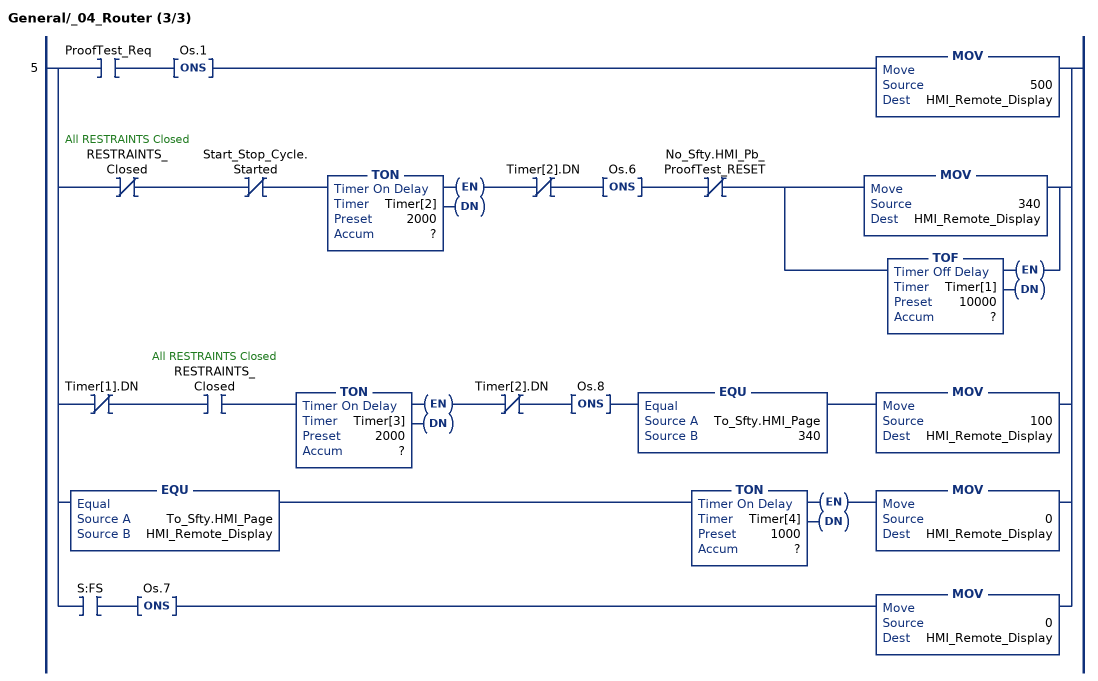
   5: [XIC(ProofTest_Req) ONS(Os.1) MOV(500,HMI_Remote_Display) ,XIO(RESTRAINTS_Closed) XIO(Start_Stop_Cycle.Started) TON(Timer[2],?,?) XIO(Timer[2].DN) ONS(Os.6) XIO(No_Sfty.HMI_Pb_ProofTest_RESET) [MOV(340,HMI_Remote_Display) ,TOF(Timer[1],?,?) ] ,XIO(Timer[1].DN) XIC(RESTRAINTS_Closed) TON(Timer[3],?,?) XIO(Timer[2].DN) ONS(Os.8) EQU(To_Sfty.HMI_Page,340) MOV(100,HMI_Remote_Display) ,EQU(To_Sfty.HMI_Page,HMI_Remote_Display) TON(Timer[4],?,?) MOV(0,HMI_Remote_Display) ,XIC(S:FS) ONS(Os.7) MOV(0,HMI_Remote_Display) ];
END_ROUTINE

ROUTINE _05_Miscellany   (* ladder *)
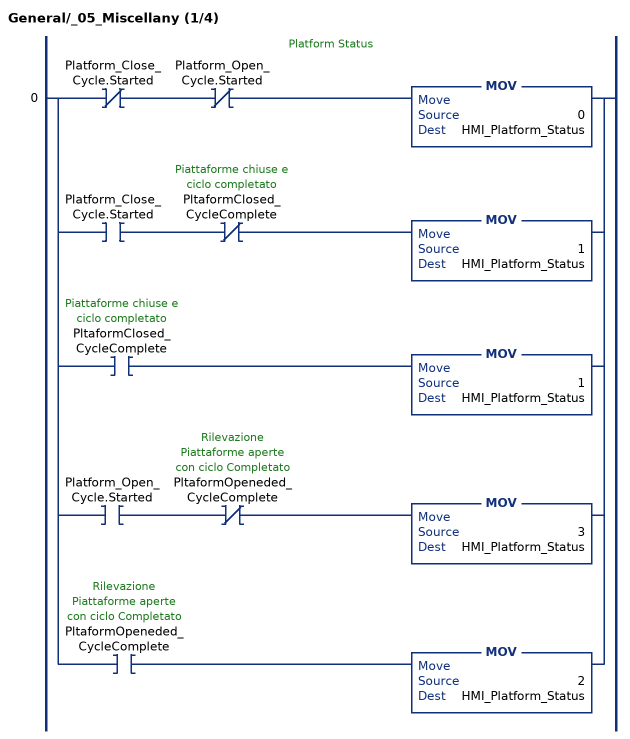
   // Platform Status
   0: [XIO(Platform_Close_Cycle.Started) XIO(Platform_Open_Cycle.Started) MOV(0,HMI_Platform_Status) ,XIC(Platform_Close_Cycle.Started) XIO(PltaformClosed_CycleComplete) MOV(1,HMI_Platform_Status) ,XIC(PltaformClosed_CycleComplete) MOV(1,HMI_Platform_Status) ,XIC(Platform_Open_Cycle.Started) XIO(PltaformOpeneded_CycleComplete) MOV(3,HMI_Platform_Status) ,XIC(PltaformOpeneded_CycleComplete) MOV(2,HMI_Platform_Status) ];
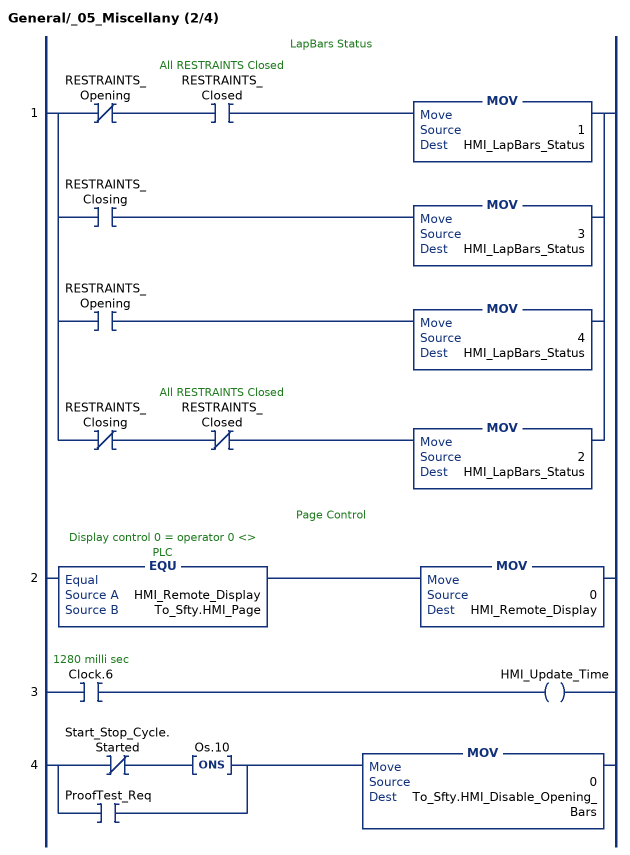
   // LapBars Status
   1: [XIO(RESTRAINTS_Opening) XIC(RESTRAINTS_Closed) MOV(1,HMI_LapBars_Status) ,XIC(RESTRAINTS_Closing) MOV(3,HMI_LapBars_Status) ,XIC(RESTRAINTS_Opening) MOV(4,HMI_LapBars_Status) ,XIO(RESTRAINTS_Closing) XIO(RESTRAINTS_Closed) MOV(2,HMI_LapBars_Status) ];
   // Page Control
   2: EQU(HMI_Remote_Display,To_Sfty.HMI_Page)MOV(0,HMI_Remote_Display);
   3: XIC(Clock.6)OTE(HMI_Update_Time);
   4: [XIO(Start_Stop_Cycle.Started) ONS(Os.10) ,XIC(ProofTest_Req) ]MOV(0,To_Sfty.HMI_Disable_Opening_Bars);
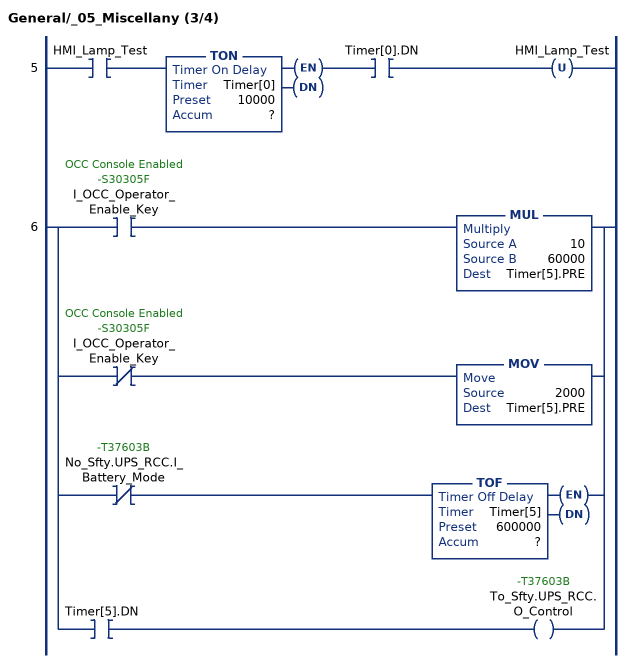
   5: XIC(HMI_Lamp_Test)TON(Timer[0],?,?)XIC(Timer[0].DN)OTU(HMI_Lamp_Test);
   6: [XIC(I_OCC_Operator_Enable_Key) MUL(10,60000,Timer[5].PRE) ,XIO(I_OCC_Operator_Enable_Key) MOV(2000,Timer[5].PRE) ,XIO(No_Sfty.UPS_RCC.I_Battery_Mode) TOF(Timer[5],?,?) ,XIC(Timer[5].DN) OTE(To_Sfty.UPS_RCC.O_Control) ];
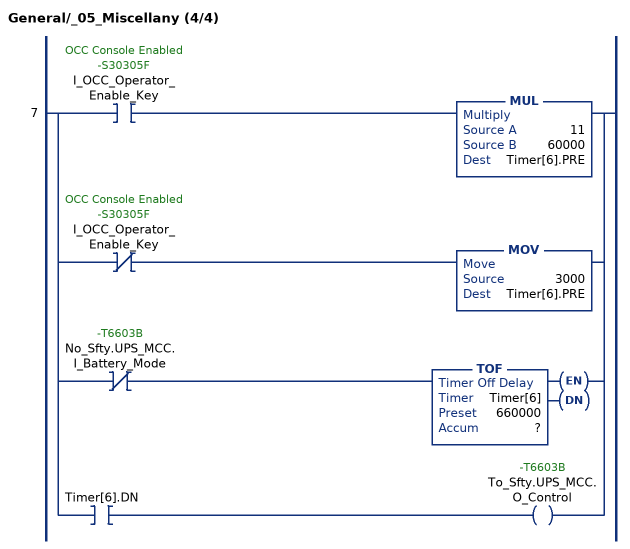
   7: [XIC(I_OCC_Operator_Enable_Key) MUL(11,60000,Timer[6].PRE) ,XIO(I_OCC_Operator_Enable_Key) MOV(3000,Timer[6].PRE) ,XIO(No_Sfty.UPS_MCC.I_Battery_Mode) TOF(Timer[6],?,?) ,XIC(Timer[6].DN) OTE(To_Sfty.UPS_MCC.O_Control) ];
END_ROUTINE

ROUTINE _06_HMI_Angle_Conversion   (* function block diagram *)
   SHEET 1
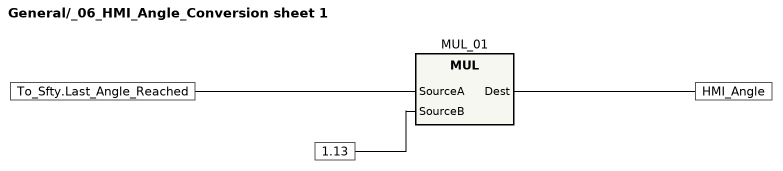
   MUL_01 : MUL(SourceA := To_Sfty.Last_Angle_Reached, SourceB := 1.13);
   HMI_Angle := MUL_01.Dest;
END_ROUTINE

ROUTINE _99_Statistics   (* ladder *)
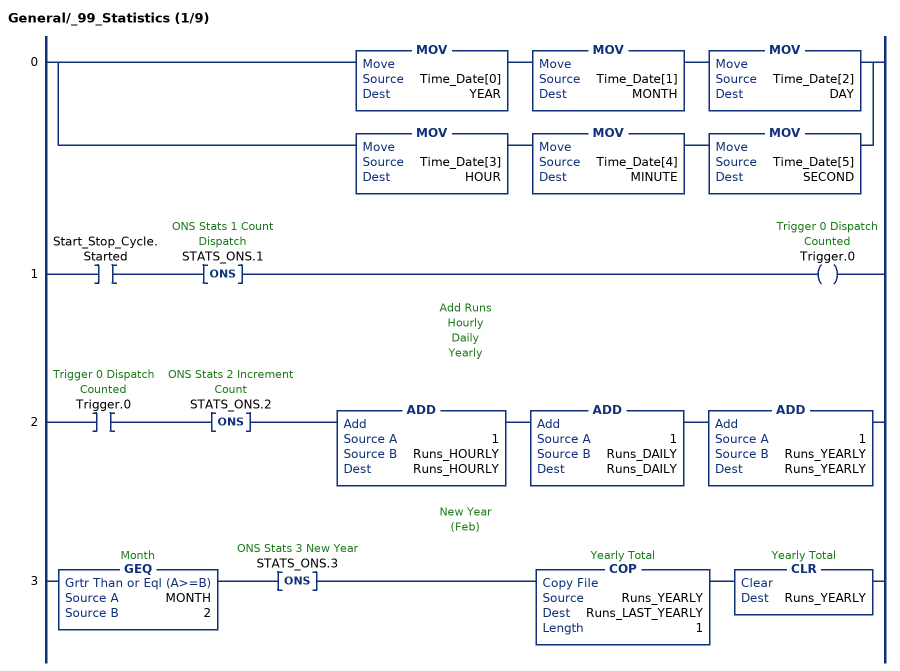
   0: [MOV(Time_Date[0],YEAR) MOV(Time_Date[1],MONTH) MOV(Time_Date[2],DAY) ,MOV(Time_Date[3],HOUR) MOV(Time_Date[4],MINUTE) MOV(Time_Date[5],SECOND) ];
   1: XIC(Start_Stop_Cycle.Started)ONS(STATS_ONS.1)OTE(Trigger.0);
   // Add Runs
   // Hourly
   // Daily
   // Yearly
   2: XIC(Trigger.0)ONS(STATS_ONS.2)ADD(1,Runs_HOURLY,Runs_HOURLY)ADD(1,Runs_DAILY,Runs_DAILY)ADD(1,Runs_YEARLY,Runs_YEARLY);
   // New Year
   // (Feb)
   3: GEQ(MONTH,2)ONS(STATS_ONS.3)COP(Runs_YEARLY,Runs_LAST_YEARLY,1)CLR(Runs_YEARLY);
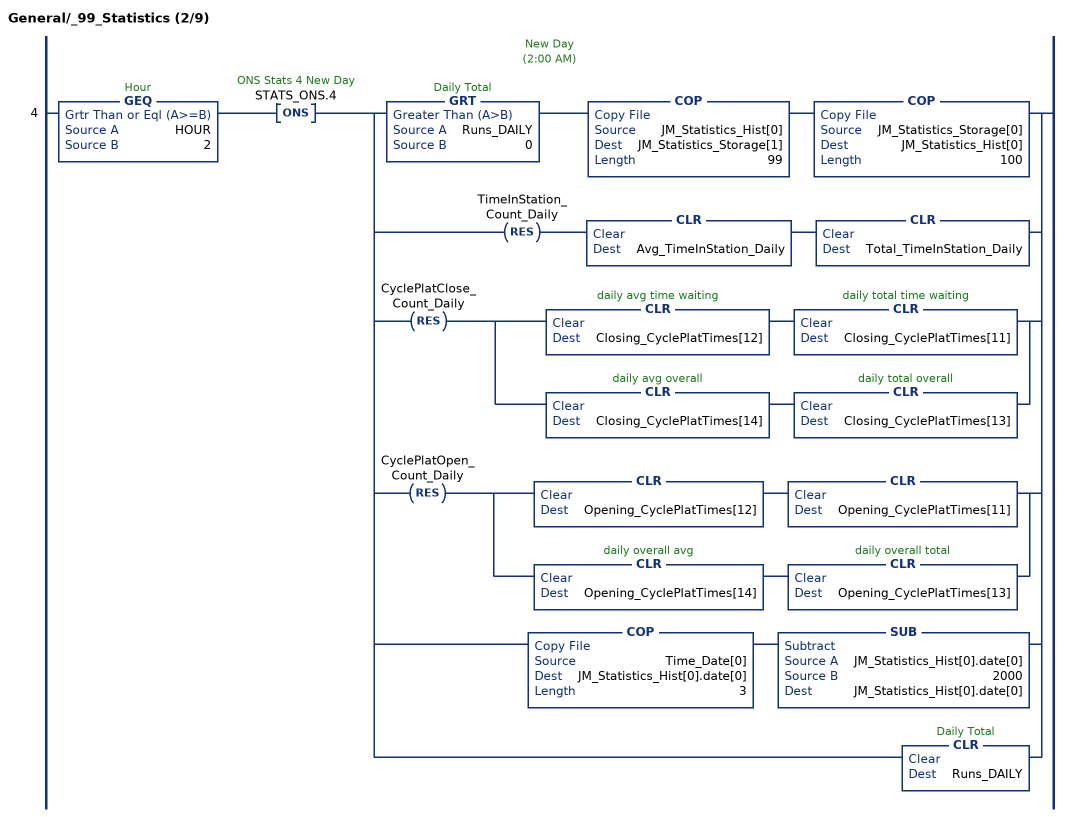
   // New Day
   // (2:00 AM)
   4: GEQ(HOUR,2)ONS(STATS_ONS.4)[[GRT(Runs_DAILY,0) COP(JM_Statistics_Hist[0],JM_Statistics_Storage[1],99) COP(JM_Statistics_Storage[0],JM_Statistics_Hist[0],100) ,RES(TimeInStation_Count_Daily) CLR(Avg_TimeInStation_Daily) CLR(Total_TimeInStation_Daily) ,RES(CyclePlatClose_Count_Daily) [CLR(Closing_CyclePlatTimes[12]) CLR(Closing_CyclePlatTimes[11]) ,CLR(Closing_CyclePlatTimes[14]) CLR(Closing_CyclePlatTimes[13]) ] ,RES(CyclePlatOpen_Count_Daily) [CLR(Opening_CyclePlatTimes[12]) CLR(Opening_CyclePlatTimes[11]) ,CLR(Opening_CyclePlatTimes[14]) CLR(Opening_CyclePlatTimes[13]) ] ,COP(Time_Date[0],JM_Statistics_Hist[0].date[0],3) SUB(JM_Statistics_Hist[0].date[0],2000,JM_Statistics_Hist[0].date[0]) ] ,CLR(Runs_DAILY) ];
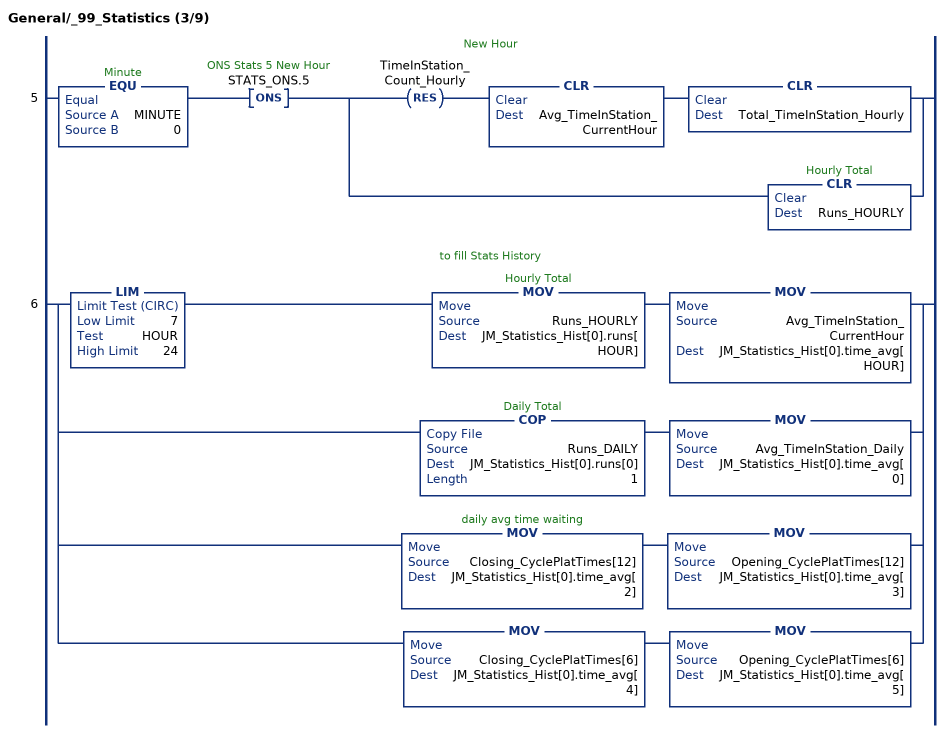
   // New Hour
   5: EQU(MINUTE,0)ONS(STATS_ONS.5)[RES(TimeInStation_Count_Hourly) CLR(Avg_TimeInStation_CurrentHour) CLR(Total_TimeInStation_Hourly) ,CLR(Runs_HOURLY) ];
   // to fill Stats History
   6: [LIM(7,HOUR,24) MOV(Runs_HOURLY,JM_Statistics_Hist[0].runs[HOUR]) MOV(Avg_TimeInStation_CurrentHour,JM_Statistics_Hist[0].time_avg[HOUR]) ,COP(Runs_DAILY,JM_Statistics_Hist[0].runs[0],1) MOV(Avg_TimeInStation_Daily,JM_Statistics_Hist[0].time_avg[0]) ,[MOV(Closing_CyclePlatTimes[12],JM_Statistics_Hist[0].time_avg[2]) MOV(Opening_CyclePlatTimes[12],JM_Statistics_Hist[0].time_avg[3]) ,MOV(Closing_CyclePlatTimes[6],JM_Statistics_Hist[0].time_avg[4]) MOV(Opening_CyclePlatTimes[6],JM_Statistics_Hist[0].time_avg[5]) ] ];
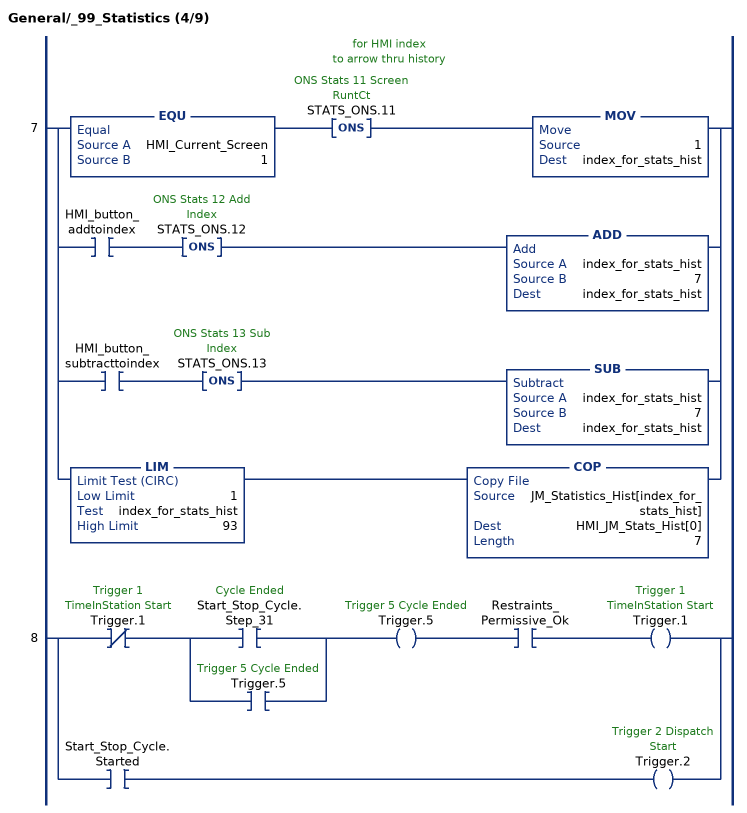
   // for HMI index
   // to arrow thru history
   7: [EQU(HMI_Current_Screen,1) ONS(STATS_ONS.11) MOV(1,index_for_stats_hist) ,[XIC(HMI_button_addtoindex) ONS(STATS_ONS.12) ADD(index_for_stats_hist,7,index_for_stats_hist) ,XIC(HMI_button_subtracttoindex) ONS(STATS_ONS.13) SUB(index_for_stats_hist,7,index_for_stats_hist) ] ,LIM(1,index_for_stats_hist,93) COP(JM_Statistics_Hist[index_for_stats_hist],HMI_JM_Stats_Hist[0],7) ];
   8: [XIO(Trigger.1) [XIC(Start_Stop_Cycle.Step_31) ,XIC(Trigger.5) ] OTE(Trigger.5) XIC(Restraints_Permissive_Ok) OTE(Trigger.1) ,XIC(Start_Stop_Cycle.Started) OTE(Trigger.2) ];
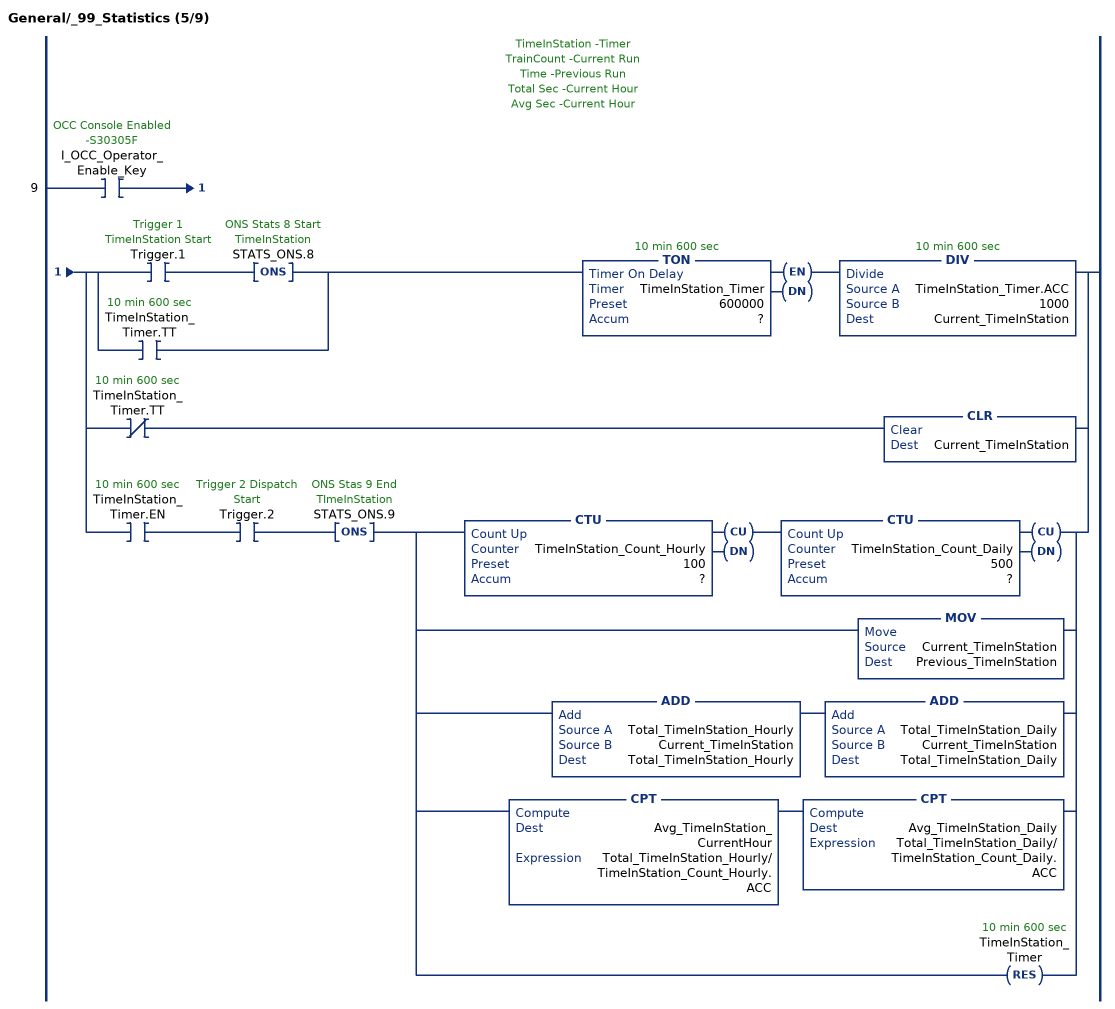
   // TimeInStation -Timer
   // TrainCount -Current Run
   // Time -Previous Run
   // Total Sec -Current Hour
   // Avg Sec -Current Hour
   9: XIC(I_OCC_Operator_Enable_Key)[[XIC(Trigger.1) ONS(STATS_ONS.8) ,XIC(TimeInStation_Timer.TT) ] TON(TimeInStation_Timer,?,?) DIV(TimeInStation_Timer.ACC,1000,Current_TimeInStation) ,XIO(TimeInStation_Timer.TT) CLR(Current_TimeInStation) ,XIC(TimeInStation_Timer.EN) XIC(Trigger.2) ONS(STATS_ONS.9) [CTU(TimeInStation_Count_Hourly,?,?) CTU(TimeInStation_Count_Daily,?,?) ,MOV(Current_TimeInStation,Previous_TimeInStation) ,ADD(Total_TimeInStation_Hourly,Current_TimeInStation,Total_TimeInStation_Hourly) ADD(Total_TimeInStation_Daily,Current_TimeInStation,Total_TimeInStation_Daily) ,CPT(Avg_TimeInStation_CurrentHour,Total_TimeInStation_Hourly/TimeInStation_Count_Hourly.ACC) CPT(Avg_TimeInStation_Daily,Total_TimeInStation_Daily/TimeInStation_Count_Daily.ACC) ,RES(TimeInStation_Timer) ] ];
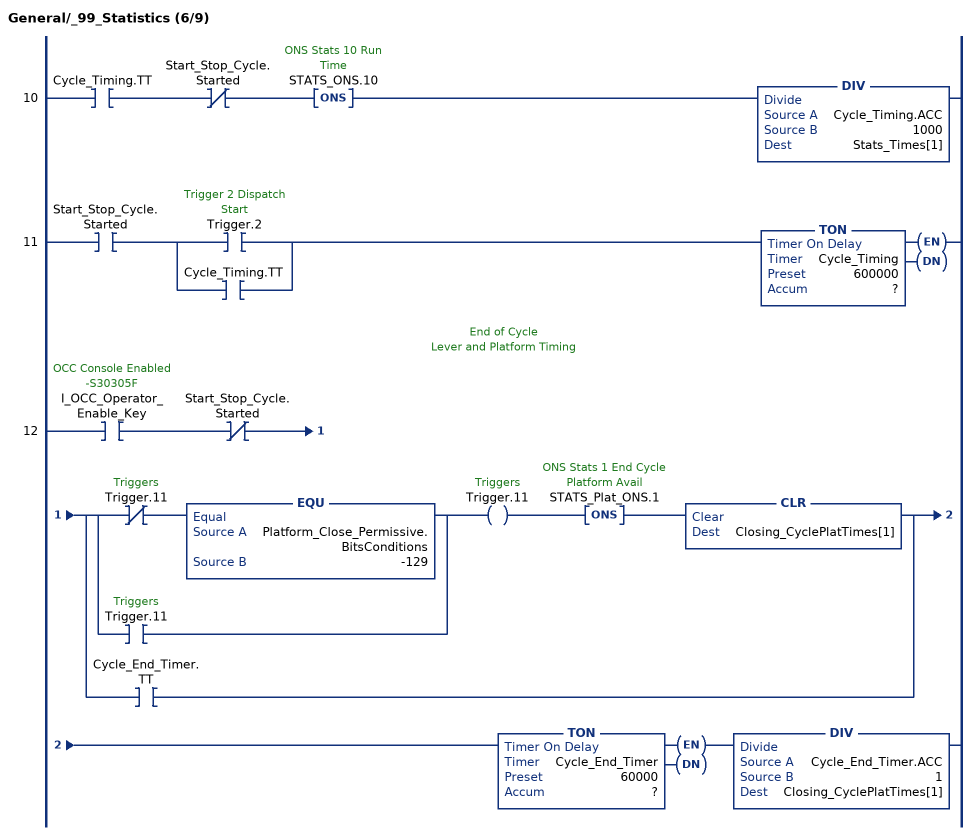
   10: XIC(Cycle_Timing.TT)XIO(Start_Stop_Cycle.Started)ONS(STATS_ONS.10)DIV(Cycle_Timing.ACC,1000,Stats_Times[1]);
   11: XIC(Start_Stop_Cycle.Started)[XIC(Trigger.2) ,XIC(Cycle_Timing.TT) ]TON(Cycle_Timing,?,?);
   // End of Cycle
   // Lever and Platform Timing
   12: XIC(I_OCC_Operator_Enable_Key)XIO(Start_Stop_Cycle.Started)[[XIO(Trigger.11) EQU(Platform_Close_Permissive.BitsConditions,-129) ,XIC(Trigger.11) ] OTE(Trigger.11) ONS(STATS_Plat_ONS.1) CLR(Closing_CyclePlatTimes[1]) ,XIC(Cycle_End_Timer.TT) ]TON(Cycle_End_Timer,?,?)DIV(Cycle_End_Timer.ACC,1,Closing_CyclePlatTimes[1]);
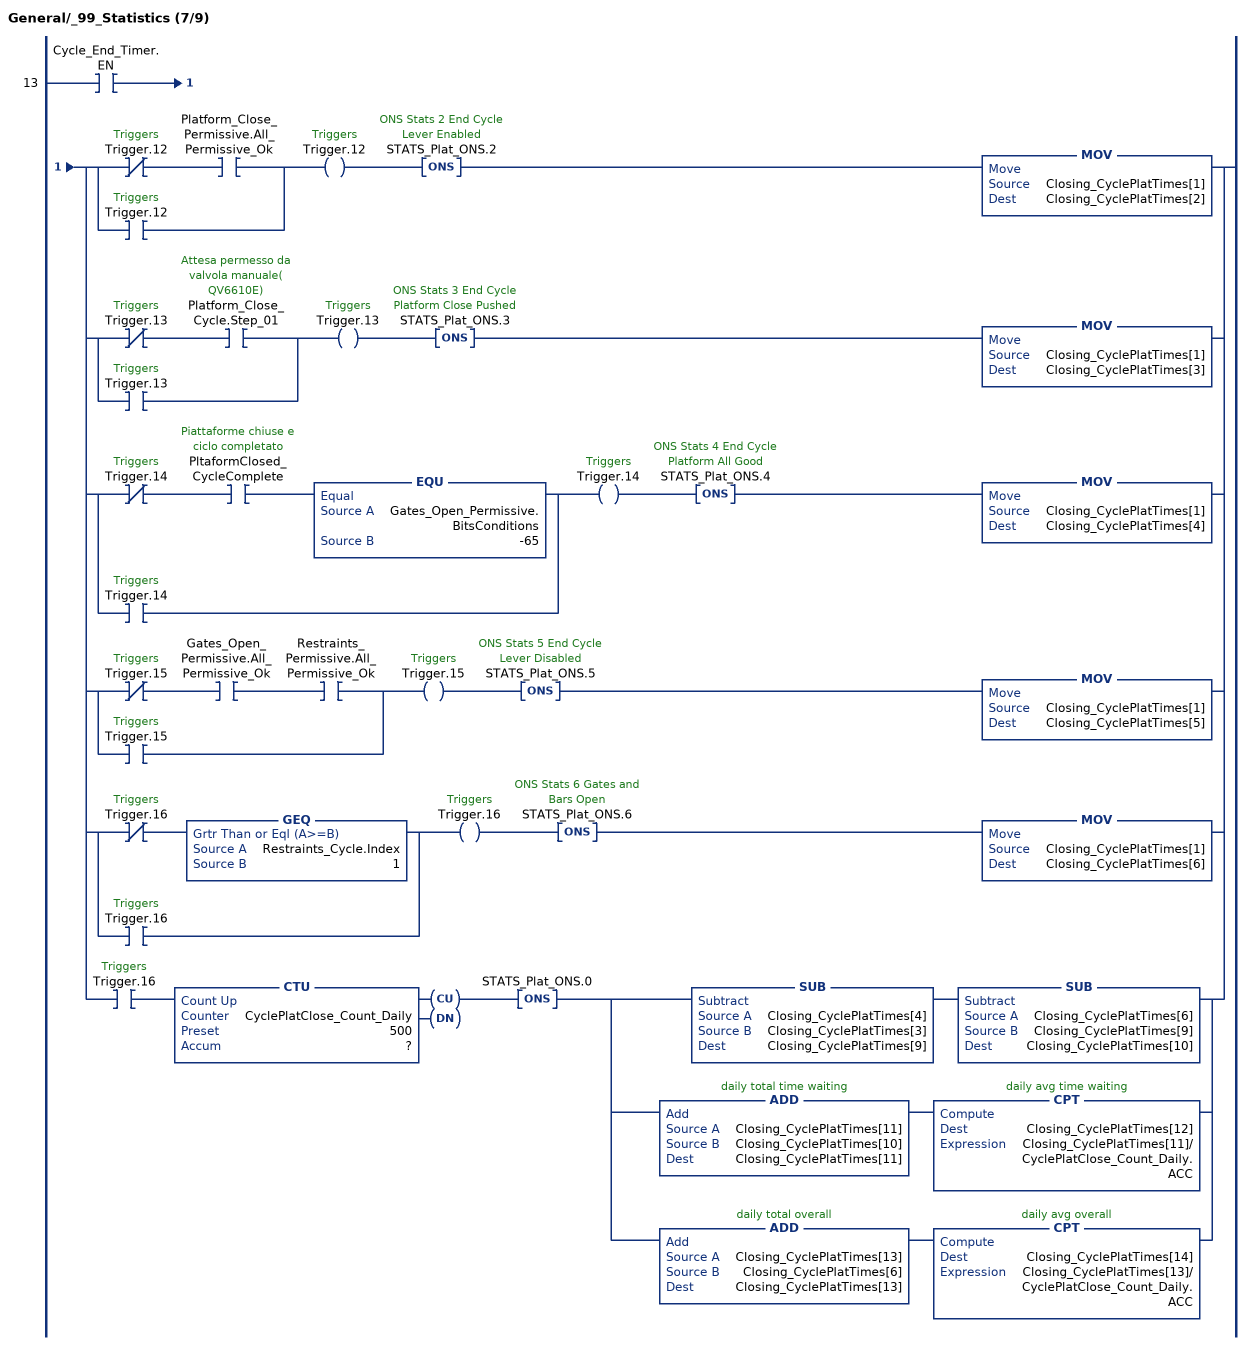
   13: XIC(Cycle_End_Timer.EN)[[XIO(Trigger.12) XIC(Platform_Close_Permissive.All_Permissive_Ok) ,XIC(Trigger.12) ] OTE(Trigger.12) ONS(STATS_Plat_ONS.2) MOV(Closing_CyclePlatTimes[1],Closing_CyclePlatTimes[2]) ,[XIO(Trigger.13) XIC(Platform_Close_Cycle.Step_01) ,XIC(Trigger.13) ] OTE(Trigger.13) ONS(STATS_Plat_ONS.3) MOV(Closing_CyclePlatTimes[1],Closing_CyclePlatTimes[3]) ,[XIO(Trigger.14) XIC(PltaformClosed_CycleComplete) EQU(Gates_Open_Permissive.BitsConditions,-65) ,XIC(Trigger.14) ] OTE(Trigger.14) ONS(STATS_Plat_ONS.4) MOV(Closing_CyclePlatTimes[1],Closing_CyclePlatTimes[4]) ,[XIO(Trigger.15) XIC(Gates_Open_Permissive.All_Permissive_Ok) XIC(Restraints_Permissive.All_Permissive_Ok) ,XIC(Trigger.15) ] OTE(Trigger.15) ONS(STATS_Plat_ONS.5) MOV(Closing_CyclePlatTimes[1],Closing_CyclePlatTimes[5]) ,[XIO(Trigger.16) GEQ(Restraints_Cycle.Index,1) ,XIC(Trigger.16) ] OTE(Trigger.16) ONS(STATS_Plat_ONS.6) MOV(Closing_CyclePlatTimes[1],Closing_CyclePlatTimes[6]) ,XIC(Trigger.16) CTU(CyclePlatClose_Count_Daily,?,?) ONS(STATS_Plat_ONS.0) [SUB(Closing_CyclePlatTimes[4],Closing_CyclePlatTimes[3],Closing_CyclePlatTimes[9]) SUB(Closing_CyclePlatTimes[6],Closing_CyclePlatTimes[9],Closing_CyclePlatTimes[10]) ,ADD(Closing_CyclePlatTimes[11],Closing_CyclePlatTimes[10],Closing_CyclePlatTimes[11]) CPT(Closing_CyclePlatTimes[12],Closing_CyclePlatTimes[11]/CyclePlatClose_Count_Daily.ACC) ,ADD(Closing_CyclePlatTimes[13],Closing_CyclePlatTimes[6],Closing_CyclePlatTimes[13]) CPT(Closing_CyclePlatTimes[14],Closing_CyclePlatTimes[13]/CyclePlatClose_Count_Daily.ACC) ] ];
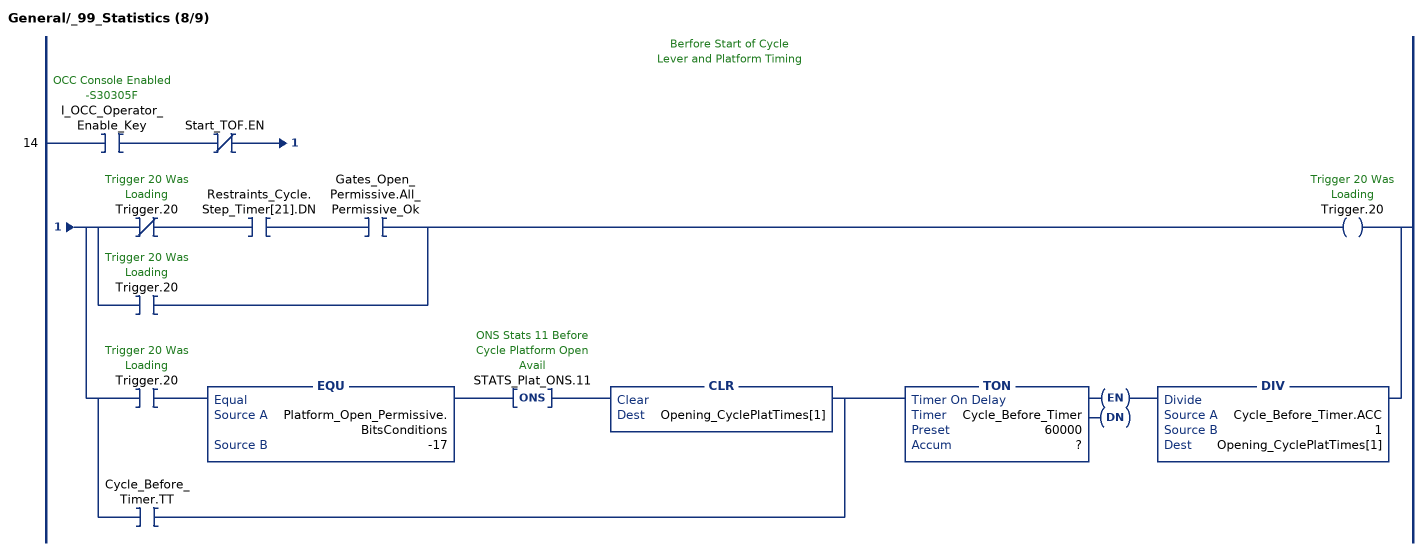
   // Berfore Start of Cycle
   // Lever and Platform Timing
   14: XIC(I_OCC_Operator_Enable_Key)XIO(Start_TOF.EN)[[XIO(Trigger.20) XIC(Restraints_Cycle.Step_Timer[21].DN) XIC(Gates_Open_Permissive.All_Permissive_Ok) ,XIC(Trigger.20) ] OTE(Trigger.20) ,[XIC(Trigger.20) EQU(Platform_Open_Permissive.BitsConditions,-17) ONS(STATS_Plat_ONS.11) CLR(Opening_CyclePlatTimes[1]) ,XIC(Cycle_Before_Timer.TT) ] TON(Cycle_Before_Timer,?,?) DIV(Cycle_Before_Timer.ACC,1,Opening_CyclePlatTimes[1]) ];
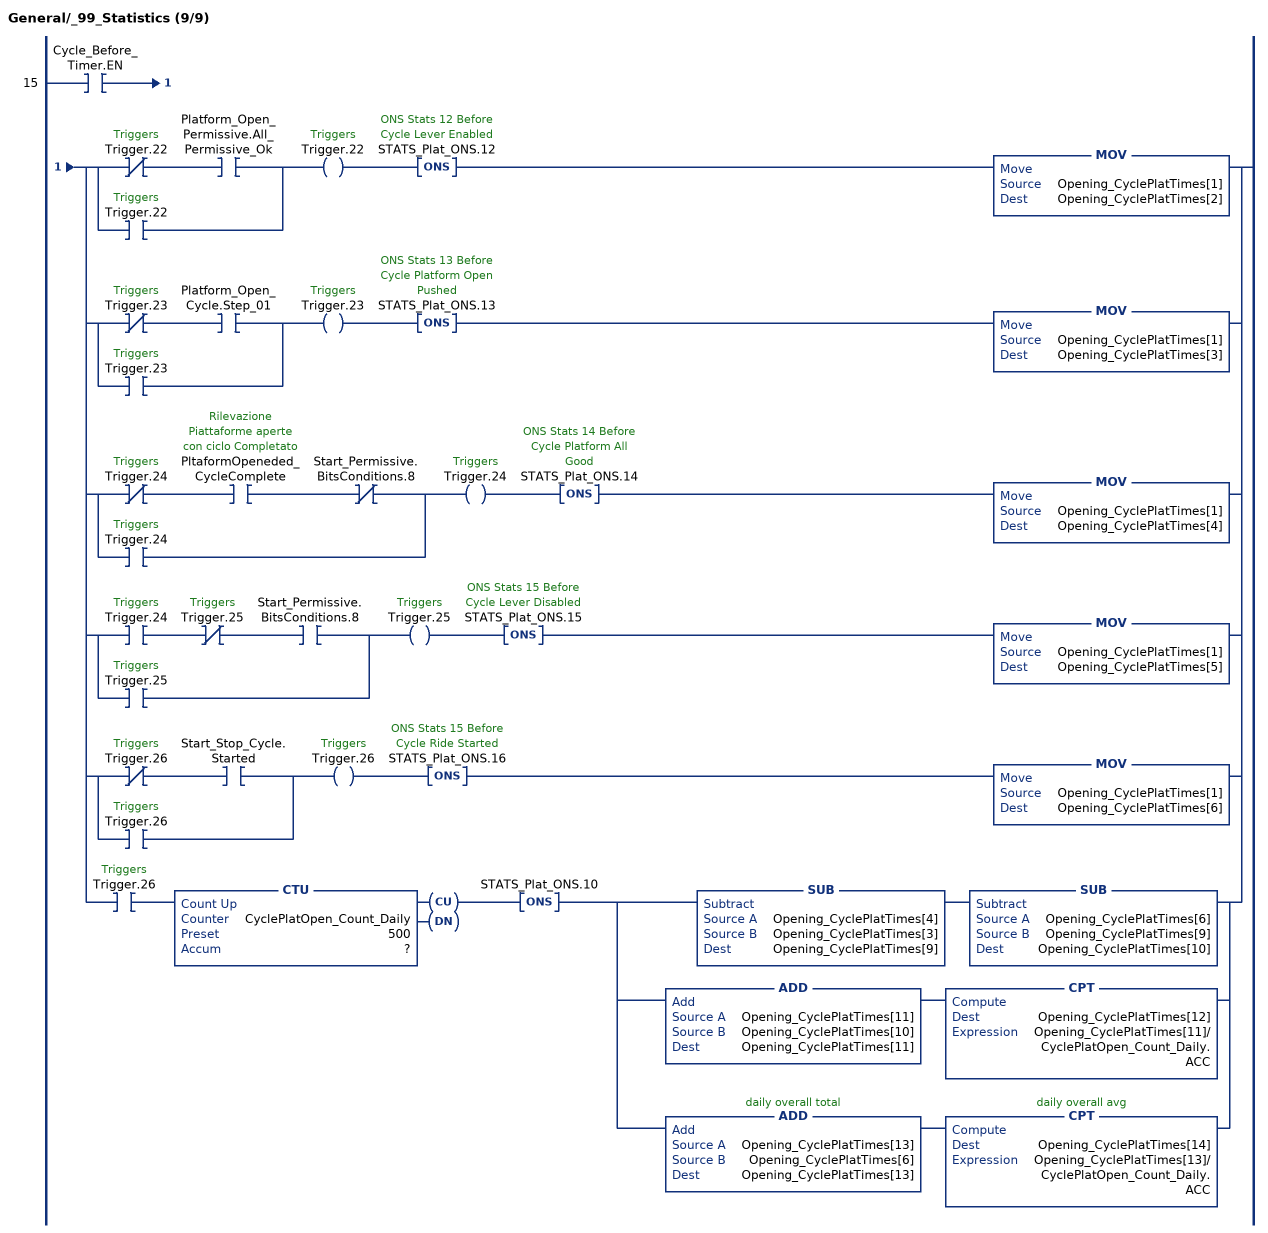
   15: XIC(Cycle_Before_Timer.EN)[[XIO(Trigger.22) XIC(Platform_Open_Permissive.All_Permissive_Ok) ,XIC(Trigger.22) ] OTE(Trigger.22) ONS(STATS_Plat_ONS.12) MOV(Opening_CyclePlatTimes[1],Opening_CyclePlatTimes[2]) ,[XIO(Trigger.23) XIC(Platform_Open_Cycle.Step_01) ,XIC(Trigger.23) ] OTE(Trigger.23) ONS(STATS_Plat_ONS.13) MOV(Opening_CyclePlatTimes[1],Opening_CyclePlatTimes[3]) ,[XIO(Trigger.24) XIC(PltaformOpeneded_CycleComplete) XIO(Start_Permissive.BitsConditions.8) ,XIC(Trigger.24) ] OTE(Trigger.24) ONS(STATS_Plat_ONS.14) MOV(Opening_CyclePlatTimes[1],Opening_CyclePlatTimes[4]) ,[XIC(Trigger.24) XIO(Trigger.25) XIC(Start_Permissive.BitsConditions.8) ,XIC(Trigger.25) ] OTE(Trigger.25) ONS(STATS_Plat_ONS.15) MOV(Opening_CyclePlatTimes[1],Opening_CyclePlatTimes[5]) ,[XIO(Trigger.26) XIC(Start_Stop_Cycle.Started) ,XIC(Trigger.26) ] OTE(Trigger.26) ONS(STATS_Plat_ONS.16) MOV(Opening_CyclePlatTimes[1],Opening_CyclePlatTimes[6]) ,XIC(Trigger.26) CTU(CyclePlatOpen_Count_Daily,?,?) ONS(STATS_Plat_ONS.10) [SUB(Opening_CyclePlatTimes[4],Opening_CyclePlatTimes[3],Opening_CyclePlatTimes[9]) SUB(Opening_CyclePlatTimes[6],Opening_CyclePlatTimes[9],Opening_CyclePlatTimes[10]) ,[ADD(Opening_CyclePlatTimes[11],Opening_CyclePlatTimes[10],Opening_CyclePlatTimes[11]) CPT(Opening_CyclePlatTimes[12],Opening_CyclePlatTimes[11]/CyclePlatOpen_Count_Daily.ACC) ,ADD(Opening_CyclePlatTimes[13],Opening_CyclePlatTimes[6],Opening_CyclePlatTimes[13]) CPT(Opening_CyclePlatTimes[14],Opening_CyclePlatTimes[13]/CyclePlatOpen_Count_Daily.ACC) ] ] ];
END_ROUTINE
